   //=============================================================================
   // START DIAGNOSTICS EVALUATION
   //=============================================================================

   //=============================================================================
   // EXISTING DEVICES
   //=============================================================================
   #tempRetValDeviceStates := DeviceStates(LADDR := #ioSystemHwId,
                                           MODE := #MODE_EXIST,
                                           STATE := #statExistingDevices);

   // Check if the block call was successful
   IF (#tempRetValDeviceStates = 0)
   THEN
       // Call ok 
       ;
   ELSIF ((#tempRetValDeviceStates = #ERR_HWID_NOT_EXISTENT)
       OR (#tempRetValDeviceStates = #ERR_LADDR_ADDRESS))
   THEN
       #ioSystemData.error := TRUE;
       #statStatus := INT_TO_WORD(#tempRetValDeviceStates);
       #statStatusID := #ID_DEVICE_STATES_EXISTING;
       #statError := TRUE;
   ELSE
       // Error handling
       #statStatus := INT_TO_WORD(#tempRetValDeviceStates);
       #statStatusID := #ID_DEVICE_STATES_EXISTING;
       #statError := TRUE;
   END_IF;

   //=============================================================================
   // FAULTY DEVICES
   //=============================================================================
   #tempRetValDeviceStates := DeviceStates(LADDR := #ioSystemHwId,
                                           MODE := #MODE_FAULTY,
                                           STATE := #statFaultyDevices);

   // Check if the block call was successful
   IF (#tempRetValDeviceStates = 0)
   THEN
       // Call ok
       ;
   ELSIF ((#tempRetValDeviceStates = #ERR_HWID_NOT_EXISTENT)
       OR (#tempRetValDeviceStates = #ERR_LADDR_ADDRESS))
   THEN
       #ioSystemData.error := TRUE;
       #statStatus := INT_TO_WORD(#tempRetValDeviceStates);
       #statStatusID := #ID_DEVICE_STATES_FAULTY;
       #statError := TRUE;
   ELSE
       // Error handling
       #statStatus := INT_TO_WORD(#tempRetValDeviceStates);
       #statStatusID := #ID_DEVICE_STATES_FAULTY;
       #statError := TRUE;
   END_IF;

   //=============================================================================
   // DISABLED DEVICES
   //=============================================================================
   #tempRetValDeviceStates := DeviceStates(LADDR := #ioSystemHwId,
                                           MODE := #MODE_DISABLED,
                                           STATE := #statDisabledDevices);

   // Check if the block call was successful
   IF (#tempRetValDeviceStates = 0)
   THEN
       // Call ok
       ;
   ELSIF ((#tempRetValDeviceStates = #ERR_HWID_NOT_EXISTENT)
       OR (#tempRetValDeviceStates = #ERR_LADDR_ADDRESS))
   THEN
       #ioSystemData.error := TRUE;
       #statStatus := INT_TO_WORD(#tempRetValDeviceStates);
       #statStatusID := #ID_DEVICE_STATES_DISABLED;
       #statError := TRUE;
   ELSE
       // Error handling
       #statStatus := INT_TO_WORD(#tempRetValDeviceStates);
       #statStatusID := #ID_DEVICE_STATES_DISABLED;
       #statError := TRUE;
   END_IF;

   //=============================================================================
   // PROBLEM DEVICES
   //=============================================================================
   #tempRetValDeviceStates := DeviceStates(LADDR := #ioSystemHwId,
                                           MODE := #MODE_PROBLEM,
                                           STATE := #statProblemDevices);

   // Check if the block call was successful
   IF (#tempRetValDeviceStates = 0)
   THEN
       // Call ok
       ;
   ELSIF ((#tempRetValDeviceStates = #ERR_HWID_NOT_EXISTENT)
       OR (#tempRetValDeviceStates = #ERR_LADDR_ADDRESS))
   THEN
       #ioSystemData.error := TRUE;
       #statStatus := INT_TO_WORD(#tempRetValDeviceStates);
       #statStatusID := #ID_DEVICE_STATES_PROBLEM;
       #statError := TRUE;
   ELSE
       // Error handling
       #statStatus := INT_TO_WORD(#tempRetValDeviceStates);
       #statStatusID := #ID_DEVICE_STATES_PROBLEM;
       #statError := TRUE;
   END_IF;

   //=============================================================================
   // Go through configured devices and check for error
   //=============================================================================
   // Initialize the pointer for the first run 
   #tempDeviceIndex := #ioSystemData.firstDevice;

   WHILE ((#tempDeviceIndex <= "USERDIAG_DEVICES_PER_IO_SYSTEM_UPPER_LIM")
       AND (#tempDeviceIndex > 0))
   DO

       IF (#ioSystemData.devices[#tempDeviceIndex].configured = TRUE)
       THEN

           IF (#statDisabledDevices[#tempDeviceIndex] = TRUE)
           THEN
               //===================
               // Device is disabled
               //===================
               #ioSystemData.devices[#tempDeviceIndex].disabled := TRUE;
               #ioSystemData.devices[#tempDeviceIndex].error := FALSE;
               #ioSystemData.devices[#tempDeviceIndex].faulty := FALSE;
               #ioSystemData.devices[#tempDeviceIndex].problem := FALSE;
               #ioSystemData.devices[#tempDeviceIndex].state := #STATE_DISABLED;

           ELSE
               #ioSystemData.devices[#tempDeviceIndex].disabled := FALSE;

               IF (#statExistingDevices[#tempDeviceIndex] = TRUE)
               THEN
                   #ioSystemData.devices[#tempDeviceIndex].exists := TRUE;

                   CASE #ioSystemData.devices[#tempDeviceIndex].state OF
                       #STATE_WAS_FAULT,
                       #STATE_WAS_LOST,
                       #STATE_WAS_DISABLED,
                       #STATE_PROBLEM_GONE:
                           ;
                       #STATE_FAULT:
                           #ioSystemData.devices[#tempDeviceIndex].state := #STATE_WAS_FAULT;
                       #STATE_LOST_CON:
                           #ioSystemData.devices[#tempDeviceIndex].state := #STATE_WAS_LOST;
                       #STATE_DISABLED:
                           #ioSystemData.devices[#tempDeviceIndex].state := #STATE_WAS_DISABLED;
                       #STATE_PROBLEM:
                           #ioSystemData.devices[#tempDeviceIndex].state := #STATE_PROBLEM_GONE;
                       ELSE
                           #ioSystemData.devices[#tempDeviceIndex].state := #STATE_OK;
                   END_CASE;

               ELSE
                   // Device not existent
                   #ioSystemData.devices[#tempDeviceIndex].error := TRUE;
                   #ioSystemData.error := TRUE;
                   #ioSystemData.devices[#tempDeviceIndex].exists := FALSE;
               END_IF; // End: Device exists


               IF (#statFaultyDevices[#tempDeviceIndex] = FALSE)
               THEN
                   // Device is not faulty
                   #ioSystemData.devices[#tempDeviceIndex].error := FALSE;
                   #ioSystemData.devices[#tempDeviceIndex].faulty := FALSE;

                   IF (#statProblemDevices[#tempDeviceIndex] = FALSE)
                   THEN
                       //============================
                       // Device has no problem
                       //============================
                       #ioSystemData.devices[#tempDeviceIndex].error := FALSE;
                       #ioSystemData.devices[#tempDeviceIndex].problem := FALSE;
                   ELSE
                       //============================
                       // Device has a problem
                       //============================
                       #ioSystemData.devices[#tempDeviceIndex].error := TRUE;
                       #ioSystemData.error := TRUE;
                       #ioSystemData.devices[#tempDeviceIndex].problem := TRUE;
                       #ioSystemData.devices[#tempDeviceIndex].state := #STATE_PROBLEM;
                   END_IF;

               ELSE
                   // Device is faulty, don't matter what happened
                   #ioSystemData.devices[#tempDeviceIndex].error := TRUE;
                   #ioSystemData.error := TRUE;
                   #ioSystemData.devices[#tempDeviceIndex].faulty := TRUE;

                   IF (#statProblemDevices[#tempDeviceIndex] = FALSE)
                   THEN
                       //============================
                       // Device has no problem
                       //============================
                       #ioSystemData.devices[#tempDeviceIndex].problem := FALSE;
                   ELSE
                       //============================
                       // Device has a problem
                       //============================
                       #ioSystemData.devices[#tempDeviceIndex].problem := TRUE;
                   END_IF;

                   IF (#statExistingDevices[#tempDeviceIndex] = FALSE)
                   THEN
                       //==========================
                       // Device is lost
                       //==========================
                       #ioSystemData.devices[#tempDeviceIndex].state := #STATE_LOST_CON;
                       #ioSystemData.devices[#tempDeviceIndex].exists := FALSE;
                   ELSE
                       //==========================
                       // Device is faulty
                       //==========================
                       #ioSystemData.devices[#tempDeviceIndex].state := #STATE_FAULT;
                       #ioSystemData.devices[#tempDeviceIndex].exists := TRUE;
                   END_IF;
               END_IF; // End: // Device is not faulty

           END_IF;

           //=============================================================================
           // Set module states
           //=============================================================================
           // Check ModuleStates if device has a problem or is faulty
           IF ((#ioSystemData.devices[#tempDeviceIndex].problem = TRUE)
               OR (#ioSystemData.devices[#tempDeviceIndex].faulty = TRUE))
           THEN

               // PROBLEM MODULE
               #tempRetValModuleStates := ModuleStates(LADDR := #ioSystemData.devices[#tempDeviceIndex].hardwareId,
                                                       MODE := #MODE_PROBLEM,
                                                       STATE := #statDeviceProblemModules);

               // Check if the block call was successful
               IF (#tempRetValModuleStates = 0)
               THEN
                   // Call ok 
                   ;
               ELSIF ((#tempRetValModuleStates = #ERR_HWID_NOT_EXISTENT)
                   OR (#tempRetValModuleStates = #ERR_LADDR_ADDRESS))
               THEN
                   #ioSystemData.error := TRUE;
                   #statStatus := INT_TO_WORD(#tempRetValModuleStates);
                   #statStatusID := #ID_MODULE_STATES_PROBLEM;
                   #statError := TRUE;
               ELSE
                   // Error handling
                   #statStatus := INT_TO_WORD(#tempRetValModuleStates);
                   #statStatusID := #ID_MODULE_STATES_PROBLEM;
                   #statError := TRUE;
               END_IF;

               // FAULTY MODULE
               #tempRetValModuleStates := ModuleStates(LADDR := #ioSystemData.devices[#tempDeviceIndex].hardwareId,
                                                       MODE := #MODE_FAULTY,
                                                       STATE := #statDeviceFaultyModules);

               // Check if the block call was successful
               IF (#tempRetValModuleStates = 0)
               THEN
                   // Call ok 
                   ;
               ELSIF ((#tempRetValModuleStates = #ERR_HWID_NOT_EXISTENT)
                   OR (#tempRetValModuleStates = #ERR_LADDR_ADDRESS))
               THEN
                   #ioSystemData.error := TRUE;
                   #statStatus := INT_TO_WORD(#tempRetValModuleStates);
                   #statStatusID := #ID_MODULE_STATES_FAULTY;
                   #statError := TRUE;
               ELSE
                   // Error handling
                   #statStatus := INT_TO_WORD(#tempRetValModuleStates);
                   #statStatusID := #ID_MODULE_STATES_FAULTY;
                   #statError := TRUE;
               END_IF;

               // EXISTING MODULE
               #tempRetValModuleStates := ModuleStates(LADDR := #ioSystemData.devices[#tempDeviceIndex].hardwareId,
                                                       MODE := #MODE_EXIST,
                                                       STATE := #statDeviceExistingModules);

               // Check if the block call was successful
               IF (#tempRetValModuleStates = 0)
               THEN
                   // Call ok 
                   ;
               ELSIF ((#tempRetValModuleStates = #ERR_HWID_NOT_EXISTENT)
                   OR (#tempRetValModuleStates = #ERR_LADDR_ADDRESS))
               THEN
                   #ioSystemData.error := TRUE;
                   #statStatus := INT_TO_WORD(#tempRetValModuleStates);
                   #statStatusID := #ID_MODULE_STATES_EXISTING;
                   #statError := TRUE;
               ELSE
                   // Error handling
                   #statStatus := INT_TO_WORD(#tempRetValModuleStates);
                   #statStatusID := #ID_MODULE_STATES_EXISTING;
                   #statError := TRUE;
               END_IF;
           END_IF;


           FOR #tempSlotIndex := 0 TO "USERDIAG_SLOTS_PER_DEVICE_UPPER_LIM" DO
               IF (#ioSystemData.devices[#tempDeviceIndex].slots[#tempSlotIndex].configured = TRUE)
               THEN
                   CASE #ioSystemData.devices[#tempDeviceIndex].slots[#tempSlotIndex].state OF
                       #STATE_WAS_FAULT,
                       #STATE_WAS_LOST,
                       #STATE_WAS_DISABLED,
                       #STATE_PROBLEM_GONE:
                           ;
                       #STATE_FAULT:
                           #ioSystemData.devices[#tempDeviceIndex].slots[#tempSlotIndex].state := #STATE_WAS_FAULT;
                       #STATE_LOST_CON:
                           #ioSystemData.devices[#tempDeviceIndex].slots[#tempSlotIndex].state := #STATE_WAS_LOST;
                       #STATE_DISABLED:
                           #ioSystemData.devices[#tempDeviceIndex].slots[#tempSlotIndex].state := #STATE_WAS_DISABLED;
                       #STATE_PROBLEM:
                           #ioSystemData.devices[#tempDeviceIndex].slots[#tempSlotIndex].state := #STATE_PROBLEM_GONE;
                       ELSE
                           #ioSystemData.devices[#tempDeviceIndex].slots[#tempSlotIndex].state := #STATE_OK;
                   END_CASE;
               END_IF;
           END_FOR;

           CASE #ioSystemData.devices[#tempDeviceIndex].state OF

               #STATE_DISABLED:
                   FOR #tempSlotIndex := 0 TO "USERDIAG_SLOTS_PER_DEVICE_UPPER_LIM" DO
                       IF (#ioSystemData.devices[#tempDeviceIndex].slots[#tempSlotIndex].configured = TRUE)
                       THEN
                           //NEW: Set all configured modules of device to disabled
                           #ioSystemData.devices[#tempDeviceIndex].slots[#tempSlotIndex].disabled := TRUE;
                           #ioSystemData.devices[#tempDeviceIndex].slots[#tempSlotIndex].error := FALSE;
                           #ioSystemData.devices[#tempDeviceIndex].slots[#tempSlotIndex].faulty := FALSE;
                           #ioSystemData.devices[#tempDeviceIndex].slots[#tempSlotIndex].problem := FALSE;
                           #ioSystemData.devices[#tempDeviceIndex].slots[#tempSlotIndex].state := #STATE_DISABLED;
                       END_IF;
                   END_FOR;

               #STATE_LOST_CON:
                   // All modules are faulty when connection is lost
                   FOR #tempSlotIndex := 0 TO "USERDIAG_SLOTS_PER_DEVICE_UPPER_LIM" DO
                       IF (#ioSystemData.devices[#tempDeviceIndex].slots[#tempSlotIndex].configured = TRUE)
                       THEN
                           #ioSystemData.devices[#tempDeviceIndex].slots[#tempSlotIndex].error := TRUE;
                           #ioSystemData.devices[#tempDeviceIndex].slots[#tempSlotIndex].faulty := TRUE;
                           #ioSystemData.devices[#tempDeviceIndex].slots[#tempSlotIndex].problem := TRUE;
                           #ioSystemData.devices[#tempDeviceIndex].slots[#tempSlotIndex].exists := FALSE;
                           #ioSystemData.devices[#tempDeviceIndex].slots[#tempSlotIndex].state := #STATE_LOST_CON;
                       END_IF;
                   END_FOR;

               #STATE_FAULT,
               #STATE_PROBLEM:
                   // The device is reachable, but faulty because of an error in a
                   // subordinated system --> check the modules
                   // Store the state of the different module in the diag DB
                   FOR #tempSlotIndex := 0 TO "USERDIAG_SLOTS_PER_DEVICE_UPPER_LIM" DO
                       IF (#ioSystemData.devices[#tempDeviceIndex].slots[#tempSlotIndex].configured = TRUE)
                       THEN
                           IF (#statDeviceProblemModules[#tempSlotIndex + 1] = TRUE)
                           THEN
                               // Problem in module
                               #ioSystemData.devices[#tempDeviceIndex].slots[#tempSlotIndex].faulty := FALSE;
                               #ioSystemData.devices[#tempDeviceIndex].slots[#tempSlotIndex].error := TRUE;
                               #ioSystemData.devices[#tempDeviceIndex].slots[#tempSlotIndex].problem := TRUE;
                               #ioSystemData.devices[#tempDeviceIndex].slots[#tempSlotIndex].state := #STATE_PROBLEM;

                               IF (#statDeviceFaultyModules[#tempSlotIndex + 1] = TRUE)
                               THEN
                                   // Fault in module
                                   #ioSystemData.devices[#tempDeviceIndex].slots[#tempSlotIndex].faulty := TRUE;
                                   #ioSystemData.devices[#tempDeviceIndex].slots[#tempSlotIndex].state := #STATE_FAULT;
                               END_IF;
                           ELSE
                               #ioSystemData.devices[#tempDeviceIndex].slots[#tempSlotIndex].error := FALSE;
                               #ioSystemData.devices[#tempDeviceIndex].slots[#tempSlotIndex].problem := FALSE;
                               #ioSystemData.devices[#tempDeviceIndex].slots[#tempSlotIndex].faulty := FALSE;
                           END_IF;

                           IF (#statDeviceExistingModules[#tempSlotIndex + 1] = TRUE)
                           THEN
                               // Module exists
                               #ioSystemData.devices[#tempDeviceIndex].slots[#tempSlotIndex].exists := TRUE;
                           ELSE
                               // Module does not exist
                               #ioSystemData.devices[#tempDeviceIndex].slots[#tempSlotIndex].exists := FALSE;
                           END_IF;
                       END_IF;
                   END_FOR;
               ELSE
                   // All modules are okay
                   FOR #tempSlotIndex := 0 TO "USERDIAG_SLOTS_PER_DEVICE_UPPER_LIM" DO
                       IF (#ioSystemData.devices[#tempDeviceIndex].slots[#tempSlotIndex].configured = TRUE)
                       THEN
                           #ioSystemData.devices[#tempDeviceIndex].slots[#tempSlotIndex].error := FALSE;
                           #ioSystemData.devices[#tempDeviceIndex].slots[#tempSlotIndex].problem := FALSE;
                           #ioSystemData.devices[#tempDeviceIndex].slots[#tempSlotIndex].faulty := FALSE;
                           #ioSystemData.devices[#tempDeviceIndex].slots[#tempSlotIndex].exists := TRUE;
                       END_IF;
                   END_FOR;
           END_CASE;
       END_IF;

       // Initialize the pointer for the next run
       #tempDeviceIndex := #ioSystemData.devices[#tempDeviceIndex].nextDevice;
   END_WHILE;


   // Write static values to outputs
   #error := #statError;
   #status := #statStatus;
   #statusID := #statStatusID;
END_FUNCTION_BLOCK

// folder: Utilities

FUNCTION "Time to WString" : WString   // FC2, SCL
{ S7_Optimized_Access := 'TRUE' }
VERSION : 0.1
   VAR_INPUT
      "Time" : Time;
   END_VAR
   VAR_TEMP
      "Time as DInt" : DInt;
      "Hours 10s Place" : DInt;
      "Hours 1s Place" : DInt;
      "Minutes 10s Place" : DInt;
      "Minutes 1s Place" : DInt;
      "Seconds 10s Place" : DInt;
      "Seconds 1s Place" : DInt;
      "Time Elements" : Array[0..4] of WString;
      Length : Int;
      "String Box" : WString;
      "DInt Box" : DInt;
   END_VAR
   VAR CONSTANT
      "Milliseconds per 10 Hours" : DInt := 36000000;
      "Milliseconds per Hour" : DInt := 3600000;
      "Milliseconds per 10 Minutes" : DInt := 600000;
      "Milliseconds per Minute" : DInt := 60000;
      "Milliseconds per 10 Seconds" : DInt := 10000;
      "Milliseconds per Second" : DInt := 1000;
   END_VAR
BEGIN
   REGION GET INPUT
       #"Time as DInt" := #Time;
   END_REGION

   REGION CONVERT TIME INTO INDIVIDUAL PLACE VALUES
       #"Minutes 10s Place" := #"Time as DInt" / #"Milliseconds per 10 Minutes";
       #"Minutes 1s Place" := (#"Time as DInt" / #"Milliseconds per Minute") MOD 10;
       #"Seconds 10s Place" := (#"Time as DInt" MOD #"Milliseconds per Minute") / #"Milliseconds per 10 Seconds";
       #"Seconds 1s Place" := (#"Time as DInt" / #"Milliseconds per Second") MOD 10;
   END_REGION

   REGION "ADD SIGN"
       #"Time Elements"[0] := wstring#'';
       IF #"Minutes 10s Place" < 0 OR
           #"Minutes 1s Place" < 0 OR
           #"Seconds 10s Place" < 0 OR
           #"Seconds 1s Place" < 0 THEN
            #"Time Elements"[0] := wstring#'-';
       END_IF;
   END_REGION

   REGION CONVERT PLACE VALUES INTO COMPONENT STRINGS
       // MINUTES
       #"DInt Box" := #"Minutes 10s Place" * 10 + #"Minutes 1s Place";
       #"String Box" := DINT_TO_WSTRING(IN := #"DInt Box");
       #"String Box" := "Strip Sign"("WString":=#"String Box");
       #"String Box" := "Add Leading"("Leading Character" := WCHAR#'0',
                                      "Desired Length" := 2,
                                      "String" := #"String Box");
       #"Time Elements"[1] := #"String Box";
       // COLON
       #"Time Elements"[2] := WSTRING#':';
       // SECONDS
       #"DInt Box" := #"Seconds 10s Place" * 10 + #"Seconds 1s Place";
       #"String Box" := DINT_TO_WSTRING(IN := #"DInt Box");
       #"String Box" := "Strip Sign"("WString":=#"String Box");
       #"String Box" := "Add Leading"("Leading Character" := WCHAR#'0',
                                      "Desired Length" := 2,
                                      "String" := #"String Box");
       #"Time Elements"[3] := #"String Box";
   END_REGION


   REGION RETURN VALUE
       #"Time to WString" := CONCAT_WSTRING(IN1 := #"Time Elements"[0],
                                            IN2 := #"Time Elements"[1],
                                            IN3 := #"Time Elements"[2],
                                            IN4 := #"Time Elements"[3]);
   END_REGION
END_FUNCTION

FUNCTION "Strip Sign" : WString   // FC3, SCL
{ S7_Optimized_Access := 'TRUE' }
VERSION : 0.1
   VAR_INPUT
      WString : WString;
   END_VAR
   VAR_TEMP
      Length : Int;
      "String Box" : WString;
      "Test Character" : WString;
   END_VAR
   VAR CONSTANT
      "+" : WChar := WCHAR#'+';
      "-" : WChar := WCHAR#'-';
   END_VAR
BEGIN
   #"String Box" := #WString;
   #"Test Character" := LEFT_WSTRING(IN := #"String Box",
                                     L := 1);
   IF #"Test Character" = #"+" OR #"Test Character" = #"-" THEN
       #Length := LEN(#"String Box");
       #"String Box" := RIGHT_WSTRING(IN := #"String Box", L := #Length - 1);

   END_IF;
   #"Strip Sign" := #"String Box";
END_FUNCTION

FUNCTION "WString to Time" : Time   // FC10, SCL
{ S7_Optimized_Access := 'TRUE' }
VERSION : 0.1
   VAR_INPUT
      WString : WString;
   END_VAR
   VAR_TEMP
      Count : UInt;
      "DInt Box" : DInt;
      "String Box" : WString [5];
      "Time Box" : Time;
      "WChar Array" : Array[0..4] of WChar;
   END_VAR
   VAR CONSTANT
      "ms/(10 hr)" : DInt := 36000000;
      "ms/hr" : DInt := 3600000;
      "ms/(10 min)" : DInt := 600000;
      "ms/min" : DInt := 60000;
      "ms/(10 sec)" : DInt := 10000;
      "ms/sec" : DInt := 1000;
   END_VAR
BEGIN
   REGION EXPLODE INPUT

       #"String Box" := #WString;
       IF #"String Box" = WSTRING#'' THEN
           #"String Box" := WSTRING#'00:00';
       END_IF;

       Strg_TO_Chars(Strg := #"String Box",
                     pChars := 0,
                     Cnt => #Count,
                     Chars := #"WChar Array");

   END_REGION

   REGION CONVERT ARRAY ELEMENTS TO TIME

       // 10S OF MINUTES
       #"DInt Box" := WCHAR_TO_DINT(IN := #"WChar Array"[0]) - 16#30;
       #"Time Box" := #"Time Box" + #"DInt Box" * #"ms/(10 min)";

       // MINUTES
       #"DInt Box" := WCHAR_TO_DINT(IN := #"WChar Array"[1]) - 16#30;
       #"Time Box" := #"Time Box" + #"DInt Box" * #"ms/min";

       // 10S OF SECONDS
       #"DInt Box" := WCHAR_TO_DINT(IN := #"WChar Array"[3]) - 16#30;
       #"Time Box" := #"Time Box" + #"DInt Box" * #"ms/(10 sec)";

       // SECONDS
       #"DInt Box" := WCHAR_TO_DINT(IN := #"WChar Array"[4]) - 16#30;
       #"Time Box" := #"Time Box" + #"DInt Box" * #"ms/sec";

   END_REGION


   REGION RETURN VALUE

       #"WString to Time" := #"Time Box";

   END_REGION
END_FUNCTION

FUNCTION "WString Timer to Real" : Real   // FC13, SCL
{ S7_Optimized_Access := 'TRUE' }
VERSION : 0.1
   VAR_INPUT
      wstring : WString;
   END_VAR
   VAR CONSTANT
      msPerSec : Real := 1000.0;
   END_VAR
BEGIN
   #"WString Timer to Real" := DINT_TO_REAL(TIME_TO_DINT("WString to Time"(#wstring))) / #msPerSec;
END_FUNCTION

FUNCTION "Word Wrap" : WString   // FC28, SCL
{ S7_Optimized_Access := 'TRUE' }
VERSION : 0.1
   VAR_INPUT
      stringIn : WString;
      maxLength : Int;
   END_VAR
   VAR_TEMP
      length : Int;
      charBox : Array[0.."lStringLen"] of WChar;
      stringBox : Array[0.."lStringLen"] of WString["lStringLen"];
      count : UInt;
      status : Int;
      i : Int;
      pStringBox : Int;
      output : WString;
      savedOutput : WString;
      lineBox : Array[0..10] of WString["lStringLen"];
      pLineBox : Int;
      lengthTest : WString;
   END_VAR
   VAR CONSTANT
      space : WString := WSTRING#' ';
      blank : WString;
      lineBreak : WString := WSTRING#'$L';
   END_VAR
BEGIN
   #length := LEN(#stringIn);

   IF #length <= #maxLength THEN
       #output := #stringIn;
   END_IF;

   IF #length > #maxLength THEN

       Strg_TO_Chars(
                     Strg := #stringIn,
                     pChars := 0,
                     Cnt => #count,
                     Chars := #charBox
       );

       FOR #i := 0 TO "lStringLen" DO

           IF #charBox[#i] = #space THEN
               IF #charBox[#i + 1] = #space THEN
                   EXIT;
               END_IF;
           END_IF;

           IF #i = 0 THEN
               #stringBox[#pStringBox] := #charBox[#i];
           END_IF;

           IF #i >= 1 THEN
               #stringBox[#pStringBox] := CONCAT_WSTRING(IN1 := #stringBox[#pStringBox],
                                                         IN2 := #charBox[#i]);
           END_IF;

           IF #charBox[#i] = #space THEN
               #stringBox[#pStringBox] := "Trim"(#stringBox[#pStringBox]);
               #pStringBox := #pStringBox + 1;
           END_IF;

           IF #charBox[#i] = #lineBreak THEN
               #stringBox[#pStringBox] := LEFT(IN := #stringBox[#pStringBox],
                                               L := LEN(#stringBox[#pStringBox]) - 1);
               #pStringBox := #pStringBox + 1;
               #stringBox[#pStringBox] := #lineBreak;
               #pStringBox := #pStringBox + 1;
           END_IF;

       END_FOR;


       FOR #i := 0 TO "lStringLen" DO

           IF #stringBox[#i] = #blank THEN
               IF #stringBox[#i + 1] = #blank THEN
                   #lineBox[#pLineBox] := "Trim"(#lineBox[#pLineBox]);
                   EXIT;
               END_IF;
           END_IF;

           IF #stringBox[#i] = #lineBreak THEN
               #lineBox[#pLineBox] := "Trim"(#lineBox[#pLineBox]);
               #pLineBox := #pLineBox + 1;
               #lineBox[#pLineBox] := #lineBreak;
               #pLineBox := #pLineBox + 1;
           END_IF;


           IF #stringBox[#i] <> #lineBreak THEN

               IF #i = 0 THEN
                   #lengthTest := #stringBox[#i];
               END_IF;

               IF #i >= 1 THEN
                   #lengthTest := CONCAT_WSTRING(IN1 := #lineBox[#pLineBox],
                                                 IN2 := #space,
                                                 IN3 := #stringBox[#i]);
               END_IF;

               IF LEN(#lengthTest) <= #maxLength THEN
                   #lineBox[#pLineBox] := #lengthTest;
               END_IF;

               IF LEN(#lengthTest) > #maxLength THEN
                   #lineBox[#pLineBox] := "Trim"(#lineBox[#pLineBox]);
                   #lineBox[#pLineBox] := "Trim"(#lineBox[#pLineBox]);
                   #pLineBox := #pLineBox + 1;
                   #lineBox[#pLineBox] := #stringBox[#i];
               END_IF;
           END_IF;

       END_FOR;

       FOR #i := 0 TO 10 DO

           IF #lineBox[#i] = #space OR #lineBox[#i] = WString#'' THEN
               EXIT;
           END_IF;
           IF #i = 0 THEN
               #output := #lineBox[#i];
           END_IF;
           IF #i >= 1 THEN
               IF #lineBox[#i] = #lineBreak THEN
                   #output := #output;
               END_IF;
               IF #lineBox[#i] <> #lineBreak THEN
                   #output := CONCAT_WSTRING(IN1 := #output,
                                             IN2 := #lineBreak,
                                             IN3 := #lineBox[#i]);
               END_IF;
           END_IF;

       END_FOR;

       #output := "Trim"(#output);

   END_IF;

   #"Word Wrap" := #output;
END_FUNCTION

FUNCTION "Trim" : WString   // FC29, SCL
{ S7_Optimized_Access := 'TRUE' }
VERSION : 0.1
   VAR_INPUT
      stringIn : WString;
   END_VAR
   VAR_TEMP
      output : WString;
   END_VAR
   VAR CONSTANT
      space : WString := WSTRING#' ';
   END_VAR
BEGIN
   #output := #stringIn;
   IF LEFT(IN := #output, L := 1) = #space THEN
       #output := RIGHT(IN := #output, L := LEN(#output) - 1);
   END_IF;
   IF RIGHT(IN := #output, L := 1) = #space THEN
       #output := LEFT(IN := #output, L := LEN(#output) - 1);
   END_IF;
   #Trim := #output;
END_FUNCTION

// ===== library types =====

TYPE "Table Row Data"
   STRUCT
      address : UInt;
      ordered : Bool;
      pbSelection : Struct
         actuate : Bool;
         animate : USInt;
      END_STRUCT;
      rtBackground : Struct
         animate : USInt;
      END_STRUCT;
      tfDropZone : Struct
         animate : USInt;
         value : WString[20];
      END_STRUCT;
      tfLine : Struct
         animate : USInt;
         value : WString[20];
      END_STRUCT;
      tfPartNumber : Struct
         animateDL : USInt;
         animateSL : USInt;
         value : WString[40];
      END_STRUCT;
      tfTime : Struct
         animate : USInt;
         value : WString[20];
      END_STRUCT;
   END_STRUCT;
END_TYPE

TYPE "Station Assignment: Button Details Data"
   STRUCT
      alloted : Struct
         animate : USInt;
         value : WString[10];
      END_STRUCT;
      critical : Struct
         animate : USInt;
         value : WString[10];
      END_STRUCT;
      label : Struct
         animate : USInt;
         value : WString[2];
      END_STRUCT;
      partNumber : Struct
         animate : USInt;
         value : WString[40];
      END_STRUCT;
      select : Struct
         actuate : Bool;
         animate : USInt;
      END_STRUCT;
   END_STRUCT;
END_TYPE

(* ===== HMI "HMI_RT_1" =====
system functions are stored by id; their names below are inferred from use
connection "Main HMI": ETHERNET, S7_1500_OMS

HMI tags "Default tag table"
   "Clock_Byte" : Byte = PLC Clock_Byte AT %MB0, 100 ms
   "HMI_screenNumber" : Int = PLC HMI.screenNumber AT %DB1.DBW0, 100 ms
   "HMI_barcode" : Barcode Screen = PLC HMI.barcode AT %DB1.DBW0, 100 ms
   "HMI_partCall_row{0}" : Table Row = PLC HMI.partCall.row[0], 100 ms
   "HMI_partCall_row{1}" : Table Row = PLC HMI.partCall.row[1], 100 ms
   "HMI_partCall_row{2}" : Table Row = PLC HMI.partCall.row[2], 100 ms
   "HMI_partCall_row{3}" : Table Row = PLC HMI.partCall.row[3], 100 ms
   "HMI_partCall_row{4}" : Table Row = PLC HMI.partCall.row[4], 100 ms
   "HMI_partCall_row{5}" : Table Row = PLC HMI.partCall.row[5], 100 ms
   "HMI_partCall_row{6}" : Table Row = PLC HMI.partCall.row[6], 100 ms
   "HMI_partCall_row{7}" : Table Row = PLC HMI.partCall.row[7], 100 ms
   "HMI_partCall_row{8}" : Table Row = PLC HMI.partCall.row[8], 100 ms
   "HMI_partCall_row{9}" : Table Row = PLC HMI.partCall.row[9], 100 ms
   "HMI_partCall_row{10}" : Table Row = PLC HMI.partCall.row[10], 100 ms
   "HMI_settings_stations_selectBtns{0}" : PB Data: Text Label = PLC HMI.settings.stations.selectBtns[0], 100 ms
   "HMI_settings_stations_selectBtns{1}" : PB Data: Text Label = PLC HMI.settings.stations.selectBtns[1], 100 ms
   "HMI_settings_stations_selectBtns{2}" : PB Data: Text Label = PLC HMI.settings.stations.selectBtns[2], 100 ms
   "HMI_settings_stations_selectBtns{3}" : PB Data: Text Label = PLC HMI.settings.stations.selectBtns[3], 100 ms
   "HMI_settings_stations_selectBtns{4}" : PB Data: Text Label = PLC HMI.settings.stations.selectBtns[4], 100 ms
   "HMI_settings_stations_selectBtns{5}" : PB Data: Text Label = PLC HMI.settings.stations.selectBtns[5], 100 ms
   "HMI_settings_stations_selectBtns{6}" : PB Data: Text Label = PLC HMI.settings.stations.selectBtns[6], 100 ms
   "HMI_settings_stations_selectBtns{7}" : PB Data: Text Label = PLC HMI.settings.stations.selectBtns[7], 100 ms
   "HMI_settings_stations_selectBtns{8}" : PB Data: Text Label = PLC HMI.settings.stations.selectBtns[8], 100 ms
   "HMI_settings_stations_selectBtns{9}" : PB Data: Text Label = PLC HMI.settings.stations.selectBtns[9], 100 ms
   "HMI_settings_stations_selectBtns{10}" : PB Data: Text Label = PLC HMI.settings.stations.selectBtns[10], 100 ms
   "HMI_settings_stations_selectBtns{11}" : PB Data: Text Label = PLC HMI.settings.stations.selectBtns[11], 100 ms
   "HMI_settings_kp8_buttons{0}" : PB Data: Text Label = PLC HMI.settings.kp8.buttons[0], 100 ms
   "HMI_settings_kp8_buttons{7}" : PB Data: Text Label = PLC HMI.settings.kp8.buttons[7], 100 ms
   "HMI_settings_kp8_buttons{3}" : PB Data: Text Label = PLC HMI.settings.kp8.buttons[3], 100 ms
   "HMI_settings_kp8_buttons{6}" : PB Data: Text Label = PLC HMI.settings.kp8.buttons[6], 100 ms
   "HMI_settings_kp8_buttons{2}" : PB Data: Text Label = PLC HMI.settings.kp8.buttons[2], 100 ms
   "HMI_settings_kp8_buttons{5}" : PB Data: Text Label = PLC HMI.settings.kp8.buttons[5], 100 ms
   "HMI_settings_kp8_buttons{1}" : PB Data: Text Label = PLC HMI.settings.kp8.buttons[1], 100 ms
   "HMI_settings_kp8_buttons{4}" : PB Data: Text Label = PLC HMI.settings.kp8.buttons[4], 100 ms
   "HMI_settings_stations_selCount" : Int = PLC HMI.settings.stations.selCount, 100 ms
   "HMI_settings_viewingStation_btns{0}" : Station Assignment: Button Details = PLC HMI.settings.viewingStation.btns[0], 100 ms
   "HMI_settings_viewingStation_btns{1}" : Station Assignment: Button Details = PLC HMI.settings.viewingStation.btns[1], 100 ms
   "HMI_settings_viewingStation_btns{2}" : Station Assignment: Button Details = PLC HMI.settings.viewingStation.btns[2], 100 ms
   "HMI_settings_viewingStation_btns{3}" : Station Assignment: Button Details = PLC HMI.settings.viewingStation.btns[3], 100 ms
   "HMI_settings_viewingStation_btns{4}" : Station Assignment: Button Details = PLC HMI.settings.viewingStation.btns[4], 100 ms
   "HMI_settings_viewingStation_btns{5}" : Station Assignment: Button Details = PLC HMI.settings.viewingStation.btns[5], 100 ms
   "HMI_settings_viewingStation_previous" : PB Data: Graphic/Text List = PLC HMI.settings.viewingStation.previous, 100 ms
   "HMI_settings_viewingStation_next" : PB Data: Graphic/Text List = PLC HMI.settings.viewingStation.next, 100 ms
   "HMI_settings_stations_selectAll" : PB Data: Text Label = PLC HMI.settings.stations.selectAll, 100 ms
   "HMI_settings_partNumber_assign" : PB Data: Text Label = PLC HMI.settings.partNumber.assign, 100 ms
   "HMI_settings_partNumber_ioField" : IO Field Data: Part Number = PLC HMI.settings.partNumber.ioField, 100 ms
   "HMI_settings_alotted_assign" : PB Data: Text Label = PLC HMI.settings.alotted.assign, 100 ms
   "HMI_settings_alotted_ioField" : IO Field Data: Timers = PLC HMI.settings.alotted.ioField, 100 ms
   "HMI_settings_critical_assign" : PB Data: Text Label = PLC HMI.settings.critical.assign, 100 ms
   "HMI_settings_critical_ioField" : IO Field Data: Timers = PLC HMI.settings.critical.ioField, 100 ms
   "HMI_settings_kp8_selectButtons" : PB Data: Text Label = PLC HMI.settings.kp8.selectButtons, 100 ms
   "HMI_settings_viewingStation_dzData" : Drop Zone Data = PLC HMI.settings.viewingStation.dzData, 100 ms
   "HMI_settings_viewingStation_lineData" : Line Label Data = PLC HMI.settings.viewingStation.lineData, 100 ms
   "HMI_settings_stations_prevGroup" : PB Data: Graphic/Text List = PLC HMI.settings.stations.prevGroup, 100 ms
   "HMI_settings_stations_nextGroup" : PB Data: Graphic/Text List = PLC HMI.settings.stations.nextGroup, 100 ms
   "HMI_settings_viewingStation_name" : WString[20] = PLC HMI.settings.viewingStation.name, 100 ms
   "HMI_tableNav_top" : PB Data: Graphic/Text List = PLC HMI.tableNav.top, 100 ms
   "HMI_tableNav_pageUp" : PB Data: Graphic/Text List = PLC HMI.tableNav.pageUp, 100 ms
   "HMI_tableNav_lineUp" : PB Data: Graphic/Text List = PLC HMI.tableNav.lineUp, 100 ms
   "HMI_tableNav_lineDown" : PB Data: Graphic/Text List = PLC HMI.tableNav.lineDown, 100 ms
   "HMI_tableNav_pageDown" : PB Data: Graphic/Text List = PLC HMI.tableNav.pageDown, 100 ms
   "HMI_tableNav_bottom" : PB Data: Graphic/Text List = PLC HMI.tableNav.bottom, 100 ms
   "HMI_simStations_stations{0}" : Station Sim Data = PLC HMI.simStations.me[0] AT %DB1.DBX0.0, 100 ms
   "HMI_simStations_me{1}" : Station Sim Data = PLC HMI.simStations.me[1], 100 ms
   "HMI_simStations_me{2}" : Station Sim Data = PLC HMI.simStations.me[2], 100 ms
   "HMI_simStations_me{3}" : Station Sim Data = PLC HMI.simStations.me[3], 100 ms
   "HMI_simStations_me{4}" : Station Sim Data = PLC HMI.simStations.me[4], 100 ms
   "HMI_simStations_me{5}" : Station Sim Data = PLC HMI.simStations.me[5], 100 ms
   "HMI_simStations_me{6}" : Station Sim Data = PLC HMI.simStations.me[6], 100 ms
   "HMI_simStations_me{7}" : Station Sim Data = PLC HMI.simStations.me[7], 100 ms
   "HMI_simStations_me{8}" : Station Sim Data = PLC HMI.simStations.me[8], 100 ms
   "HMI_simStations_me{9}" : Station Sim Data = PLC HMI.simStations.me[9], 100 ms
   "HMI_simStations_me{10}" : Station Sim Data = PLC HMI.simStations.me[10], 100 ms
   "HMI_simStations_me{11}" : Station Sim Data = PLC HMI.simStations.me[11], 100 ms
   "HMI_simStations_up" : PB Data: Graphic/Text List = PLC HMI.simStations.up, 100 ms
   "HMI_simStations_down" : PB Data: Graphic/Text List = PLC HMI.simStations.down, 100 ms
   "Log Flag" : Int = PLC "Log Buffer".logFlag AT %DB1.DBW0, 100 ms
      on ChangeValue: function_abcfba0d("Log Buffer_partReq_me{0}_address"); function_abcfba0d("Log Buffer_partReq_me{0}_timeStamp"); function_abcfba0d("Log Buffer_partReq_me{0}_reqType")
   "Log Buffer_partReq_me{0}_address" : Int = PLC "Log Buffer".partReq.me[0].address, 100 ms
   "Log Buffer_partReq_me{0}_timeStamp" : DTL = PLC "Log Buffer".partReq.me[0].timeStamp, 100 ms
   "Log Buffer_partReq_me{0}_reqType" : Int = PLC "Log Buffer".partReq.me[0].reqType, 100 ms
   "HMI_networkHealth_pnioDevices{1}" : PB Data: Text Label = PLC HMI.networkHealth.pnioDevices[1], 100 ms
   "HMI_networkHealth_pnioDevices{2}" : PB Data: Text Label = PLC HMI.networkHealth.pnioDevices[2], 1 s
   "HMI_networkHealth_pnioDevices{3}" : PB Data: Text Label = PLC HMI.networkHealth.pnioDevices[3], 1 s
   "HMI_networkHealth_pnioDevices{4}" : PB Data: Text Label = PLC HMI.networkHealth.pnioDevices[4], 1 s
   "HMI_networkHealth_pnioDevices{5}" : PB Data: Text Label = PLC HMI.networkHealth.pnioDevices[5], 1 s
   "HMI_networkHealth_pnioDevices{6}" : PB Data: Text Label = PLC HMI.networkHealth.pnioDevices[6], 1 s
   "HMI_networkHealth_pnioDevices{7}" : PB Data: Text Label = PLC HMI.networkHealth.pnioDevices[7], 1 s
   "HMI_networkHealth_pnioDevices{8}" : PB Data: Text Label = PLC HMI.networkHealth.pnioDevices[8], 1 s
   "HMI_networkHealth_pnioDevices{9}" : PB Data: Text Label = PLC HMI.networkHealth.pnioDevices[9], 1 s
   "HMI_networkHealth_pnioDevices{10}" : PB Data: Text Label = PLC HMI.networkHealth.pnioDevices[10], 1 s
   "HMI_networkHealth_pnioDevices{11}" : PB Data: Text Label = PLC HMI.networkHealth.pnioDevices[11], 1 s
   "HMI_networkHealth_pnioDevices{12}" : PB Data: Text Label = PLC HMI.networkHealth.pnioDevices[12], 1 s
   "HMI_networkHealth_pnioDevices{13}" : PB Data: Text Label = PLC HMI.networkHealth.pnioDevices[13], 1 s
   "HMI_networkHealth_pnioDevices{16}" : PB Data: Text Label = PLC HMI.networkHealth.pnioDevices[16], 1 s
   "HMI_networkHealth_pnioDevices{14}" : PB Data: Text Label = PLC HMI.networkHealth.pnioDevices[14], 1 s
   "HMI_networkHealth_pnioDevices{15}" : PB Data: Text Label = PLC HMI.networkHealth.pnioDevices[15], 1 s
   "HMI_networkHealth_pnioDevices{17}" : PB Data: Text Label = PLC HMI.networkHealth.pnioDevices[17], 1 s
   "HMI_networkHealth_pnioDevices{18}" : PB Data: Text Label = PLC HMI.networkHealth.pnioDevices[18], 1 s
   "HMI_networkHealth_pnioDevices{19}" : PB Data: Text Label = PLC HMI.networkHealth.pnioDevices[19], 1 s
   "HMI_networkHealth_pnioDevices{20}" : PB Data: Text Label = PLC HMI.networkHealth.pnioDevices[20], 1 s
   "HMI_networkHealth_pnioDevices{21}" : PB Data: Text Label = PLC HMI.networkHealth.pnioDevices[21], 1 s
   "HMI_networkHealth_pnioDevices{22}" : PB Data: Text Label = PLC HMI.networkHealth.pnioDevices[22], 1 s
   "HMI_networkHealth_pnioDevices{31}" : PB Data: Text Label = PLC HMI.networkHealth.pnioDevices[31], 1 s
   "HMI_networkHealth_pnioDevices{32}" : PB Data: Text Label = PLC HMI.networkHealth.pnioDevices[32], 1 s
   "HMI_networkHealth_pnioDevices{29}" : PB Data: Text Label = PLC HMI.networkHealth.pnioDevices[29], 1 s
   "HMI_networkHealth_pnioDevices{30}" : PB Data: Text Label = PLC HMI.networkHealth.pnioDevices[30], 1 s
   "HMI_networkHealth_pnioDevices{27}" : PB Data: Text Label = PLC HMI.networkHealth.pnioDevices[27], 1 s
   "HMI_networkHealth_pnioDevices{28}" : PB Data: Text Label = PLC HMI.networkHealth.pnioDevices[28], 1 s
   "HMI_networkHealth_pnioDevices{23}" : PB Data: Text Label = PLC HMI.networkHealth.pnioDevices[23], 1 s
   "HMI_networkHealth_pnioDevices{24}" : PB Data: Text Label = PLC HMI.networkHealth.pnioDevices[24], 1 s
   "HMI_networkHealth_pnioDevices{25}" : PB Data: Text Label = PLC HMI.networkHealth.pnioDevices[25], 1 s
   "HMI_networkHealth_pnioDevices{26}" : PB Data: Text Label = PLC HMI.networkHealth.pnioDevices[26], 1 s
   "HMI_networkHealth_pnioDevices{33}" : PB Data: Text Label = PLC HMI.networkHealth.pnioDevices[33], 1 s
   "HMI_networkHealth_pnioDevices{34}" : PB Data: Text Label = PLC HMI.networkHealth.pnioDevices[34], 1 s
   "HMI_networkHealth_pnioDevices{35}" : PB Data: Text Label = PLC HMI.networkHealth.pnioDevices[35], 1 s
   "HMI_networkHealth_pnioDevices{36}" : PB Data: Text Label = PLC HMI.networkHealth.pnioDevices[36], 1 s
   "HMI_networkHealth_pnioDevices{37}" : PB Data: Text Label = PLC HMI.networkHealth.pnioDevices[37], 1 s
   "HMI_networkHealth_pnioDevices{38}" : PB Data: Text Label = PLC HMI.networkHealth.pnioDevices[38], 1 s
   "HMI_networkHealth_pnioDevices{39}" : PB Data: Text Label = PLC HMI.networkHealth.pnioDevices[39], 1 s
   "HMI_networkHealth_pnioDevices{40}" : PB Data: Text Label = PLC HMI.networkHealth.pnioDevices[40], 1 s
   "HMI_networkHealth_pnioDevices{41}" : PB Data: Text Label = PLC HMI.networkHealth.pnioDevices[41], 1 s
   "HMI_networkHealth_pnioDevices{42}" : PB Data: Text Label = PLC HMI.networkHealth.pnioDevices[42], 1 s
   "HMI_networkHealth_pnioDevices{43}" : PB Data: Text Label = PLC HMI.networkHealth.pnioDevices[43], 1 s
   "HMI_networkHealth_pnioDevices{44}" : PB Data: Text Label = PLC HMI.networkHealth.pnioDevices[44], 1 s
   "HMI_networkHealth_pnioDevices{45}" : PB Data: Text Label = PLC HMI.networkHealth.pnioDevices[45], 1 s
   "HMI_networkHealth_pnioDevices{46}" : PB Data: Text Label = PLC HMI.networkHealth.pnioDevices[46], 1 s
   "HMI_networkHealth_pnioDevices{47}" : PB Data: Text Label = PLC HMI.networkHealth.pnioDevices[47], 1 s
   "HMI_networkHealth_pnioDevices{48}" : PB Data: Text Label = PLC HMI.networkHealth.pnioDevices[48], 1 s
   "HMI_networkHealth_et200spPopUp" : Station: ET200SP Comm Debug Data = PLC HMI.networkHealth.et200spPopUp, 1 s
   "HMI_networkHealth_kp8PopUp" : Station: KP8 Comm Debug Data = PLC HMI.networkHealth.kp8PopUp, 1 s
   "HMI_networkHealth_selectedDevice" : Int = PLC HMI.networkHealth.selectedDevice, 1 s
   "EMP IDB_stations_me{0}_partNumbers{0}" : WString[40] = PLC "EMP IDB".stations.me[0].partNumbers[0], 1 s
   "EMP IDB_stations_me{0}_partNumbers{1}" : WString[40] = PLC "EMP IDB".stations.me[0].partNumbers[1], 1 s
   "EMP IDB_stations_me{0}_partNumbers{2}" : WString[40] = PLC "EMP IDB".stations.me[0].partNumbers[2], 1 s
   "EMP IDB_stations_me{0}_partNumbers{3}" : WString[40] = PLC "EMP IDB".stations.me[0].partNumbers[3], 1 s
   "EMP IDB_stations_me{0}_partNumbers{4}" : WString[40] = PLC "EMP IDB".stations.me[0].partNumbers[4], 1 s
   "EMP IDB_stations_me{0}_partNumbers{5}" : WString[40] = PLC "EMP IDB".stations.me[0].partNumbers[5], 1 s
   "EMP IDB_stations_me{0}_partNumbers{6}" : WString[40] = PLC "EMP IDB".stations.me[0].partNumbers[6], 1 s
   "EMP IDB_stations_me{0}_partNumbers{7}" : WString[40] = PLC "EMP IDB".stations.me[0].partNumbers[7], 1 s
   "EMP IDB_stations_me{1}_partNumbers{0}" : WString[40] = PLC "EMP IDB".stations.me[1].partNumbers[0], 1 s
   "EMP IDB_stations_me{1}_partNumbers{1}" : WString[40] = PLC "EMP IDB".stations.me[1].partNumbers[1], 1 s
   "EMP IDB_stations_me{1}_partNumbers{2}" : WString[40] = PLC "EMP IDB".stations.me[1].partNumbers[2], 1 s
   "EMP IDB_stations_me{1}_partNumbers{3}" : WString[40] = PLC "EMP IDB".stations.me[1].partNumbers[3], 1 s
   "EMP IDB_stations_me{1}_partNumbers{4}" : WString[40] = PLC "EMP IDB".stations.me[1].partNumbers[4], 1 s